                   IF (#tempRetValue <> 0) THEN
                     #LKinCtrl_OffsetContour.returnValue := #tempRetValue;
                     #LKinCtrl_OffsetContour."region" := #COFF_REGION_TYPE_RAD_COMP_LIN_CIRC;
                     #LKinCtrl_OffsetContour.subBlockNumber := 35052;
                     #LKinCtrl_OffsetContour.internalNumber := 333;
                     RETURN;
                   END_IF;



                 END_IF;

                 // Calculate end coordinate of "next" linear command
                 // Calculate orthogonal and tangential vector for next but one circular commamnd
                 #tempRetValue := "LKinCtrl_CalcCircTangOrthPathPlane"(circlePoint := #tempNextCmdIn.endPoint,
                                                                       circleCenterPoint := #tempNextButOneCmdIn.circleCenterPoint,
                                                                       pathPlane := #pathPlane,
                                                                       compDirection := #compensationDirection,
                                                                       pathChoice := #tempNextButOneCmdIn.pathChoice,
                                                                       vUnitTangentialPathPlane => #tempNextButOneCmdOut.tangentialUnitVecStart,
                                                                       vUnitOrthogonalPathPlane => #tempNextButOneCmdOut.orthogonalUnitVecStart);

                 IF (#tempRetValue <> 0) THEN
                   #LKinCtrl_OffsetContour.returnValue := #tempRetValue;
                   #LKinCtrl_OffsetContour."region" := #COFF_REGION_TYPE_RAD_COMP_LIN_CIRC;
                   #LKinCtrl_OffsetContour.subBlockNumber := 35056;
                   #LKinCtrl_OffsetContour.internalNumber := 334;
                   RETURN;
                 END_IF;


                 // Scale othogonal vector with tool radius to get orthogonal shift
                 #tempNextButOneCmdOut.orthogonalShiftStart := "LKinCtrl_VecScale"(vIn := #tempNextButOneCmdOut.orthogonalUnitVecStart,
                                                                                   factor := #toolRadius);

                 #tempNextButOneCmdOut.startPointOrthShifted := "LKinCtrl_VecAdd"(vIn1 := #tempNextCmdIn.endPoint,
                                                                                  vIn2 := #tempNextButOneCmdOut.orthogonalShiftStart);

                 // Calculate radius of circle
                 #tempNextCmdOut.circleRadius := "LKinCtrl_VecAbs"("LKinCtrl_VecSub"(vIn1 := #tempNextButOneCmdOut.startPointOrthShifted,
                                                                                                                                       vIn2 := #tempNextButOneCmdIn.circleCenterPoint));


                 // ########## Intersection point of 1st linear and 2nd circular command  ##########
                 #tempRetValue := "LKinCtrl_CalcLineCircleIntersectionPoint"(startPointLine := #tempNextCmdOut.endPointOrthShifted,
                                                                             endPointLine := #tempNextCmdOut.endPointOrthTangShifted,
                                                                             circleCenter := #tempNextButOneCmdIn.circleCenterPoint,
                                                                             circleRadius := #tempNextCmdOut.circleRadius,
                                                                             intersectionPointA => #tempPa,
                                                                             intersectionPointB => #tempPb);

                 IF (#tempRetValue <> 0) THEN
                   #LKinCtrl_OffsetContour.returnValue := #tempRetValue;
                   #LKinCtrl_OffsetContour."region" := #COFF_REGION_TYPE_RAD_COMP_LIN_CIRC;
                   #LKinCtrl_OffsetContour.subBlockNumber := 35061;
                   #LKinCtrl_OffsetContour.internalNumber := 335;
                   RETURN;
                 END_IF;

                 // Two intersection points, use the one which is closer to the circle start point
                 #tempDistance1 := "LKinCtrl_VecAbs"("LKinCtrl_VecSub"(vIn1 := #tempNextCmdOut.endPointOrthShifted, vIn2 := #tempPa));
                 #tempDistance2 := "LKinCtrl_VecAbs"("LKinCtrl_VecSub"(vIn1 := #tempNextCmdOut.endPointOrthShifted, vIn2 := #tempPb));

                 IF (#tempDistance1 < #tempDistance2) THEN
                   #tempNextCmdOut.endPoint := #tempPa;
                 ELSE
                   #tempNextCmdOut.endPoint := #tempPb;
                 END_IF;

               END_REGION
               // ############# N E X T   B U T   O N E   C M D  -  N O N E #############
             ELSE
               REGION Next but one command NONE
                 // V01.01.02 AW 2020-10-13
                 // Check if current end point is in opposite direction, e.g. small command length with big tool radius etc.
                 // Avoid reversal movement

                 // Calculate difference vector of uncompensated current and next end point
                 #tempDirectionUncompensatedVec := "LKinCtrl_VecSub"(vIn1 := #tempCurrentPoint, vIn2 := #tempNextCmdIn.endPoint);
                 #tempDirectionUncompensatedUnitVec := "LKinCtrl_VecUnit"(#tempDirectionUncompensatedVec);

                 // Calculate difference vector of compensated current and next end point
                 #tempDirectionCompensatedVec := "LKinCtrl_VecSub"(vIn1 := #tempCurrentPointRadComp, vIn2 := #tempNextCmdOut.endPoint);
                 #tempDirectionCompensatedUnitVec := "LKinCtrl_VecUnit"(#tempDirectionCompensatedVec);

                 // Calculate length between current compensated and next compensated end point
                 #tempLengthCompensatedPointDifferenceVec := "LKinCtrl_VecAbs"(#tempDirectionCompensatedVec);

                 // Check if vectors are parallel 
                 IF (((ABS(#tempDirectionUncompensatedUnitVec.x) - ABS(#tempDirectionCompensatedUnitVec.x)) < #COFF_TOLERANCE) AND
                   ((ABS(#tempDirectionUncompensatedUnitVec.y) - ABS(#tempDirectionCompensatedUnitVec.y)) < #COFF_TOLERANCE) AND
                   ((ABS(#tempDirectionUncompensatedUnitVec.z) - ABS(#tempDirectionCompensatedUnitVec.z)) < #COFF_TOLERANCE))
                 THEN
                   // Opposite direction?
                   IF ((ABS(#tempDirectionUncompensatedUnitVec.x + #tempDirectionCompensatedUnitVec.x) < #COFF_TOLERANCE) AND
                     (ABS(#tempDirectionUncompensatedUnitVec.y + #tempDirectionCompensatedUnitVec.y) < #COFF_TOLERANCE) AND
                     (ABS(#tempDirectionUncompensatedUnitVec.z + #tempDirectionCompensatedUnitVec.z) < #COFF_TOLERANCE))
                   THEN
                     // Throw error
                     #LKinCtrl_OffsetContour.returnValue := #ERR_COFF_LINEAR_CMD_AND_TOOL_RADIUS_LEAD_TO_REVERSAL;
                     #LKinCtrl_OffsetContour."region" := #COFF_REGION_TYPE_RAD_COMP_LIN_NONE;
                     #LKinCtrl_OffsetContour.subBlockNumber := 0;
                     #LKinCtrl_OffsetContour.internalNumber := 336;
                     RETURN;

                     // // Possible solution - NOT used!
                     // // Use tangential and orthogonal shift
                     // // Scale tangential vector with point difference (compensated points) to get tangential shift
                     // #tempNextCmdOut.tangentiaShiftEnd := "LKinCtrl_VecScale"(vIn := #tempNextCmdOut.tangentialUnitVecEnd,
                     //                                                          factor := #tempLengthCompensatedPointDifferenceVec);

                     // // Re-calculate orthogonal and (new) tangential shifted next target coordinate
                     // // next command end point will be equal to last command end point --> no reversal
                     // #tempNextCmdOut.endPointOrthTangShifted := "LKinCtrl_VecAdd"(vIn1 := #tempNextCmdOut.endPointOrthShifted,
                     //                                                              vIn2 := #tempNextCmdOut.tangentiaShiftEnd);

                     // // Use tangential and orthogonal shift - assign new value
                     // #tempNextCmdOut.endPoint := #tempNextCmdOut.endPointOrthTangShifted;

                   ELSE
                     // Same direction
                     ;// Nothing to do
                   END_IF;
                 ELSE
                   // V01.01.03
                   ;// Nothing to do
                 END_IF;

               END_REGION
             END_IF;

             REGION Additional plausibility check
               #tempRetValue := "LKinCtrl_CalcAngleBetweenVectors"(point1 := #tempNextCmdOut.endPoint,
                                                                   point2 := #tempNextCmdIn.endPoint,
                                                                   intersectionPoint := #tempCurrentPoint,
                                                                   angle => #tempAngle);

               IF (#tempRetValue <> 0) THEN
                 #LKinCtrl_OffsetContour.returnValue := #tempRetValue;
                 #LKinCtrl_OffsetContour."region" := #COFF_REGION_TYPE_RAD_COMP_LIN_GEN;
                 #LKinCtrl_OffsetContour.subBlockNumber := 35059;
                 #LKinCtrl_OffsetContour.internalNumber := 340;
                 RETURN;
               END_IF;

               IF (#tempAngle > #COFF_CIRC_REVERSAL_TOLERANCE_ANGLE)
               THEN
                 #LKinCtrl_OffsetContour.returnValue := #ERR_COFF_NO_SOLUTION_FOR_GIVEN_LINEAR_CMD;
                 #LKinCtrl_OffsetContour."region" := #COFF_REGION_TYPE_RAD_COMP_LIN_GEN;
                 #LKinCtrl_OffsetContour.subBlockNumber := 0;
                 #LKinCtrl_OffsetContour.internalNumber := 341;
                 RETURN;
               END_IF;

             END_REGION
           ELSE
             // Use radius compensated coordinates
             CASE #pathPlane OF
               "CP_XY":
                 #tempNextCmdOut.endPoint.x := #tempCurrentPointRadComp.x;
                 #tempNextCmdOut.endPoint.y := #tempCurrentPointRadComp.y;
                 #tempNextCmdOut.endPoint.z := #tempNextCmdOut.endPoint.z;

               "CP_XZ":
                 #tempNextCmdOut.endPoint.x := #tempCurrentPointRadComp.x;
                 #tempNextCmdOut.endPoint.y := #tempNextCmdOut.endPoint.y;
                 #tempNextCmdOut.endPoint.z := #tempCurrentPointRadComp.z;

               "CP_YZ":
                 #tempNextCmdOut.endPoint.x := #tempNextCmdOut.endPoint.x;
                 #tempNextCmdOut.endPoint.y := #tempCurrentPointRadComp.y;
                 #tempNextCmdOut.endPoint.z := #tempCurrentPointRadComp.z;
             END_CASE;
           END_IF;
         END_IF;
       END_REGION

       REGION Next command CIRCULAR
         // ############# N E X T   C M D  -  C I R C U L A R #############
         // ##############################################
         IF (#tempNextCmdOut.cmdType = "LKINCTRL_MC_MOVECIRCULARABS") THEN

           // Distinguish between different circular modes
           IF (#tempNextCmdIn.circleMode = "CM_BORDER") THEN

             // ------------ Via an intermediate point and the end point ("CircMode" = 0) ------------
             // Caluclate center point of circle with given start point, end point and intermediate point
             #tempRetValue := "LKinCtrl_CalcCircCenterByIntermediatePointAndEndPoint"(circleStartPoint := #tempCurrentPoint,
                                                                                      circleEndPoint := #tempNextCmdIn.endPoint,
                                                                                      circleIntermediatePoint := #tempNextCmdIn.circleIntermediatePoint,
                                                                                      pathPlane := #pathPlane,
                                                                                      circleCenterPoint => #tempNextCmdIn.circleCenterPoint);

             IF (#tempRetValue <> 0) THEN
               #LKinCtrl_OffsetContour.returnValue := #tempRetValue;
               #LKinCtrl_OffsetContour."region" := #COFF_REGION_TYPE_RAD_COMP_NEXT_CMD_CIRC;
               #LKinCtrl_OffsetContour.subBlockNumber := 35057;

               #LKinCtrl_OffsetContour.internalNumber := 401;
               RETURN;
             END_IF;

             // Calculate path choice
             #tempRetValue := "LKinCtrl_CalcCircPathChoiceByIntermediatePointAndEndPoint"(circleStartPoint := #tempCurrentPoint,
                                                                                          circleEndPoint := #tempNextCmdIn.endPoint,
                                                                                          circleintermediatePoint := #tempNextCmdIn.circleIntermediatePoint,
                                                                                          pathPlane := #pathPlane,
                                                                                          pathChoice => #tempNextCmdIn.pathChoice);

             IF (#tempRetValue <> 0) THEN
               #LKinCtrl_OffsetContour.returnValue := #tempRetValue;
               #LKinCtrl_OffsetContour."region" := #COFF_REGION_TYPE_RAD_COMP_NEXT_CMD_CIRC;
               #LKinCtrl_OffsetContour.subBlockNumber := 35058;
               #LKinCtrl_OffsetContour.internalNumber := 402;
               RETURN;
             END_IF;

           ELSIF (#tempNextCmdIn.circleMode = "CM_CENTER") THEN
             // ------------ Via the circle center and the angle in a main plane ("CircMode" = 1) ------------
             (* im oberen Teil!
             // "Third" coordinate is ignored by system - also ignore here!
             // Use start coordinate of circle instead
             IF (#pathPlane = "CP_XZ") THEN
               #tempNextCmdIn.circleCenterPoint.y := #tempCurrentPoint.y;
             ELSIF (#pathPlane = "CP_YZ") THEN
               #tempNextCmdIn.circleCenterPoint.x := #tempCurrentPoint.x;
             ELSIF (#pathPlane = "CP_XY") THEN
               #tempNextCmdIn.circleCenterPoint.z := #tempCurrentPoint.z;
             END_IF;*)
             ;

           ELSIF (#tempNextCmdIn.circleMode = "CM_RADIUS") THEN
             // ------------ Via the circle radius and the end point in a main plane ("CircMode" = 2) ------------
             // Calculate circle center point by given start / end point and radius and path choice
             #tempRetValue := "LKinCtrl_CalcCircCenterByRadiusAndEndPoint"(circleStartPoint := #tempCurrentPoint,
                                                                           circleEndPoint := #tempNextCmdIn.endPoint,
                                                                           pathPlane := #pathPlane,
                                                                           circleRadius := #tempNextCmdIn.circleRadius,
                                                                           pathChoice := #tempNextCmdIn.pathChoice,
                                                                           circCenterPoint => #tempNextCmdIn.circleCenterPoint);

             IF (#tempRetValue <> 0) THEN
               #LKinCtrl_OffsetContour.returnValue := #tempRetValue;
               #LKinCtrl_OffsetContour."region" := #COFF_REGION_TYPE_RAD_COMP_NEXT_CMD_CIRC;
               #LKinCtrl_OffsetContour.subBlockNumber := 35052;
               #LKinCtrl_OffsetContour.internalNumber := 403;
               RETURN;
             END_IF;

           END_IF;

           //REGION todo
           // 2019-03-07 - not necessary
           (*
           // ####
           // Calculate circle paramters
           #tempRetValue := "LKinCtrl_CalcCircTangOrthPathPlane"(circlePoint := #tempCurrentPoint,
                                                                 circleCenterPoint := #tempNextCmdIn.circleCenterPoint,
                                                                 pathPlane := #pathPlane,
                                                                 compDirection := #compensationDirection,
                                                                 pathChoice := #tempNextCmdIn.pathChoice,
                                                                 vUnitTangentialPathPlane => #tempNextCmdOut.tangentialUnitVecStart,
                                                                 vUnitOrthogonalPathPlane => #tempNextCmdOut.orthogonalUnitVecStart);

           IF (#tempRetValue <> 0) THEN
             #LKinCtrl_OffsetContour.returnValue := #tempRetValue;
             #LKinCtrl_OffsetContour."region" := #COFF_REGION_TYPE_RAD_COMP_LIN_CIRC;
             #LKinCtrl_OffsetContour.subBlockNumber := 35056;
             #LKinCtrl_OffsetContour.internalNumber := 404;
             RETURN;
           END_IF;

           // Scale othogonal vector with tool radius to get orthogonal shift
           #tempNextCmdOut.orthogonalShiftStart := "LKinCtrl_VecScale"(vIn := #tempNextCmdOut.orthogonalUnitVecStart,
                                                                       factor := #toolRadius);

           #tempNextCmdOut.startPointOrthShifted := "LKinCtrl_VecAdd"(vIn1 := #tempCurrentPoint,
                                                                      vIn2 := #tempNextCmdOut.orthogonalShiftStart);

           *)
           //END_REGION


           // #############  N E X T   B U T   O N E   C M D   #############
           // Check if next but one linear command has at least one component in path plane direction
           #tempRetValue := "LKinCtrl_CalcVecDistancePathPlane"(vectorInA := #tempNextCmdIn.endPoint,
                                                                vectorInB := #tempNextButOneCmdIn.endPoint,
                                                                pathPlane := #pathPlane,
                                                                distancePathPlane => #tempDistance1);

           IF (#tempRetValue <> 0) THEN
             #LKinCtrl_OffsetContour.returnValue := #tempRetValue;
             #LKinCtrl_OffsetContour."region" := #COFF_REGION_TYPE_RAD_COMP_CIRC_LIN;
             #LKinCtrl_OffsetContour.subBlockNumber := 35055;
             #LKinCtrl_OffsetContour.internalNumber := 405;
             RETURN;
           END_IF;

           // #############  N E X T   B U T   O N E   C M D   -  L I N E A R  #############
           // Linear command must have at least a motion in direction of path plane, otherwise treat as command none!
           IF (#tempNextButOneCmdOut.cmdType = "LKINCTRL_MC_MOVELINEARABS") AND (#tempDistance1 > 0.0) THEN

             REGION Next but one command LINEAR
               // 2nd linear command point 2 to point 3
               // Calculate tangential and orthogonal unit vector of direction (with respect to end point of circle)
               #tempRetValue := "LKinCtrl_CalcLineTangOrthPathPlane"(pathPlane := #pathPlane,
                                                                     compDirection := #compensationDirection,
                                                                     vInFirst := #tempNextButOneCmdIn.endPoint,
                                                                     vInSecond := #tempNextCmdIn.endPoint, // End point of circle
                                                                     vUnitTangentialPathPlane => #tempNextButOneCmdOut.tangentialUnitVecStart,
                                                                     vUnitOrthogonalPathPlane => #tempNextButOneCmdOut.orthogonalUnitVecStart);

               IF (#tempRetValue <> 0) THEN
                 #LKinCtrl_OffsetContour.returnValue := #tempRetValue;
                 #LKinCtrl_OffsetContour."region" := #COFF_REGION_TYPE_RAD_COMP_CIRC_LIN;
                 #LKinCtrl_OffsetContour.subBlockNumber := 35055;
                 #LKinCtrl_OffsetContour.internalNumber := 406;
                 RETURN;
               END_IF;

               // Scale othogonal vector with tool radius to get orthogonal shift
               #tempNextButOneCmdOut.orthogonalShiftStart := "LKinCtrl_VecScale"(vIn := #tempNextButOneCmdOut.orthogonalUnitVecStart,
                                                                                 factor := #toolRadius);

               // Scale tangential vector with tool radius to get tangential shift
               #tempNextButOneCmdOut.tangentiaShiftStart := "LKinCtrl_VecScale"(vIn := #tempNextButOneCmdOut.tangentialUnitVecStart,
                                                                                factor := #toolRadius);

               // Calculate orthogonal shifted next target coordinate
               #tempNextButOneCmdOut.startPointOrthShifted := "LKinCtrl_VecAdd"(vIn1 := #tempNextCmdIn.endPoint, // Start coordinate next but one command
                                                                                vIn2 := #tempNextButOneCmdOut.orthogonalShiftStart);

               // Calculate orthogonal and tangential shifted next target coordinate
               #tempNextButOneCmdOut.startPointOrthTangShifted := "LKinCtrl_VecAdd"(vIn1 := #tempNextButOneCmdOut.startPointOrthShifted,
                                                                                    vIn2 := #tempNextButOneCmdOut.tangentiaShiftStart);

               // ########## Intersection point of 1st circular and 2nd linear command  ##########
               // Change center point to same level with start point
               IF (#tempNextCmdIn.circleMode = "CM_BORDER") THEN
                 // ------------ Via an intermediate point and the end point ("CircMode" = 0) ------------
                 // 3D circle possible

                 // Bring circle parameter to the same level as current point
                 #tempNextCmdEndPointLevelled := #tempNextCmdIn.endPoint;
                 #tempNextCmdIntermediatePointLevelled := #tempNextCmdIn.circleIntermediatePoint;


                 // Bring coordinates to same level as current point
                 #tempNextCmdStartPointOrhtShiftLevelled := #tempCurrentPointRadComp;// #tempNextCmdOut.startPointOrthShifted;
                 #tempNextButOneStartPointOrthShiftedLevelled := #tempNextButOneCmdOut.startPointOrthShifted;
                 #tempNextButOneCmdStartPointOrthTangShiftedLevelled := #tempNextButOneCmdOut.startPointOrthTangShifted;

                 // Level parameters (third coordinate) with current point
                 CASE #pathPlane OF
                   "CP_XZ":
                     #tempNextCmdEndPointLevelled.y := #tempCurrentPoint.y;
                     #tempNextCmdIntermediatePointLevelled.y := #tempCurrentPoint.y;
                     #tempNextCmdStartPointOrhtShiftLevelled.y := #tempCurrentPoint.y;
                     #tempNextButOneStartPointOrthShiftedLevelled.y := #tempCurrentPoint.y;
                     #tempNextButOneCmdStartPointOrthTangShiftedLevelled.y := #tempCurrentPoint.y;

                   "CP_YZ":
                     #tempNextCmdEndPointLevelled.x := #tempCurrentPoint.x;
                     #tempNextCmdIntermediatePointLevelled.x := #tempCurrentPoint.x;
                     #tempNextCmdStartPointOrhtShiftLevelled.x := #tempCurrentPoint.x;
                     #tempNextButOneStartPointOrthShiftedLevelled.x := #tempCurrentPoint.x;
                     #tempNextButOneCmdStartPointOrthTangShiftedLevelled.x := #tempCurrentPoint.x;

                   "CP_XY":
                     #tempNextCmdEndPointLevelled.z := #tempCurrentPoint.z;
                     #tempNextCmdIntermediatePointLevelled.z := #tempCurrentPoint.z;
                     #tempNextCmdStartPointOrhtShiftLevelled.z := #tempCurrentPoint.z;
                     #tempNextButOneStartPointOrthShiftedLevelled.z := #tempCurrentPoint.z;
                     #tempNextButOneCmdStartPointOrthTangShiftedLevelled.z := #tempCurrentPoint.z;
                   ELSE
                     #LKinCtrl_OffsetContour.returnValue := #ERR_COFF_INTERNAL;
                     #LKinCtrl_OffsetContour."region" := #COFF_REGION_TYPE_RAD_COMP_CIRC_LIN;
                     #LKinCtrl_OffsetContour.internalNumber := 407;
                     RETURN;
                 END_CASE;

                 // Calculate new levelled circle center point
                 #tempRetValue := "LKinCtrl_CalcCircCenterByIntermediatePointAndEndPoint"(circleStartPoint := #tempCurrentPoint,
                                                                                          circleEndPoint := #tempNextCmdEndPointLevelled,
                                                                                          circleIntermediatePoint := #tempNextCmdIntermediatePointLevelled,
                                                                                          pathPlane := #pathPlane,
                                                                                          circleCenterPoint => #tempNextCmdOut.circleCenterPoint); // levelled

                 IF (#tempRetValue <> 0) THEN
                   #LKinCtrl_OffsetContour.returnValue := #tempRetValue;
                   #LKinCtrl_OffsetContour."region" := #COFF_REGION_TYPE_RAD_COMP_NEXT_CMD_CIRC;
                   #LKinCtrl_OffsetContour.subBlockNumber := 35057;
                   #LKinCtrl_OffsetContour.internalNumber := 408;
                   RETURN;
                 END_IF;

                 // Calculate modified radius - levelled
                 #tempNextCmdOut.circleRadius := "LKinCtrl_VecAbs"("LKinCtrl_VecSub"(vIn1 := #tempNextCmdStartPointOrhtShiftLevelled,
                                                                                     vIn2 := #tempNextCmdOut.circleCenterPoint));




                 #tempRetValue := "LKinCtrl_CalcLineCircleIntersectionPoint"(startPointLine := #tempNextButOneStartPointOrthShiftedLevelled,
                                                                             endPointLine := #tempNextButOneCmdStartPointOrthTangShiftedLevelled,
                                                                             circleCenter := #tempNextCmdOut.circleCenterPoint,
                                                                             circleRadius := #tempNextCmdOut.circleRadius,
                                                                             intersectionPointA => #tempPa,
                                                                             intersectionPointB => #tempPb);

                 // Relevel intersection point
                 CASE #pathPlane OF
                   "CP_XZ":
                     #tempPa.y := #tempNextCmdIn.endPoint.y;
                     #tempPb.y := #tempNextCmdIn.endPoint.y;

                   "CP_YZ":
                     #tempPa.x := #tempNextCmdIn.endPoint.x;
                     #tempPb.x := #tempNextCmdIn.endPoint.x;

                   "CP_XY":
                     #tempPa.z := #tempNextCmdIn.endPoint.z;
                     #tempPb.z := #tempNextCmdIn.endPoint.z;
                   ELSE
                     #LKinCtrl_OffsetContour.returnValue := #ERR_COFF_INTERNAL;
                     #LKinCtrl_OffsetContour."region" := #COFF_REGION_TYPE_RAD_COMP_CIRC_LIN;
                     #LKinCtrl_OffsetContour.internalNumber := 409;
                     RETURN;
                 END_CASE;

               ELSE
                 // 2D circle
                 // Calculate modified radius
                 #tempNextCmdOut.circleRadius := "LKinCtrl_VecAbs"("LKinCtrl_VecSub"(vIn1 := #tempCurrentPointRadComp,//#tempNextCmdOut.startPointOrthShifted,
                                                                                     vIn2 := #tempNextCmdIn.circleCenterPoint));

                 #tempRetValue := "LKinCtrl_CalcLineCircleIntersectionPoint"(startPointLine := #tempNextButOneCmdOut.startPointOrthShifted,
                                                                             endPointLine := #tempNextButOneCmdOut.startPointOrthTangShifted,
                                                                             circleCenter := #tempNextCmdIn.circleCenterPoint,
                                                                             circleRadius := #tempNextCmdOut.circleRadius,
                                                                             intersectionPointA => #tempPa,
                                                                             intersectionPointB => #tempPb);


               END_IF;


               IF (#tempRetValue <> 0) THEN
                 #LKinCtrl_OffsetContour.returnValue := #tempRetValue;
                 #LKinCtrl_OffsetContour."region" := #COFF_REGION_TYPE_RAD_COMP_CIRC_LIN;
                 #LKinCtrl_OffsetContour.subBlockNumber := 35061;
                 #LKinCtrl_OffsetContour.internalNumber := 410;
                 RETURN;
               END_IF;

               // Two intersection points, use the one which is closer to the circle end point
               #tempDistance1 := "LKinCtrl_VecAbs"("LKinCtrl_VecSub"(vIn1 := #tempNextCmdIn.endPoint, vIn2 := #tempPa));
               #tempDistance2 := "LKinCtrl_VecAbs"("LKinCtrl_VecSub"(vIn1 := #tempNextCmdIn.endPoint, vIn2 := #tempPb));

               IF (#tempDistance1 < #tempDistance2) THEN
                 #tempNextCmdOut.endPoint := #tempPa;
               ELSE
                 #tempNextCmdOut.endPoint := #tempPb;
               END_IF;

             END_REGION
             // #############  N E X T   B U T   O N E   C M D   -  C I R C U L A R #############
           ELSIF (#tempNextButOneCmdOut.cmdType = "LKINCTRL_MC_MOVECIRCULARABS") THEN
             REGION Next but one command CIRCULAR
               // Distinguish between different circular modes
               IF (#tempNextButOneCmdIn.circleMode = "CM_BORDER") THEN
                 // ------------ Via an intermediate point and the end point ("CircMode" = 0) ------------

                 // Caluclate center point of circle with given start point, end point and intermediate point
                 #tempRetValue := "LKinCtrl_CalcCircCenterByIntermediatePointAndEndPoint"(circleStartPoint := #tempNextCmdIn.endPoint,
                                                                                          circleEndPoint := #tempNextButOneCmdIn.endPoint,
                                                                                          circleIntermediatePoint := #tempNextButOneCmdIn.circleIntermediatePoint,
                                                                                          pathPlane := #pathPlane,
                                                                                          circleCenterPoint => #tempNextButOneCmdIn.circleCenterPoint);

                 IF (#tempRetValue <> 0) THEN
                   #LKinCtrl_OffsetContour.returnValue := #tempRetValue;
                   #LKinCtrl_OffsetContour."region" := #COFF_REGION_TYPE_RAD_COMP_CIRC_CIRC;
                   #LKinCtrl_OffsetContour.subBlockNumber := 35057;
                   #LKinCtrl_OffsetContour.internalNumber := 430;
                   RETURN;
                 END_IF;

                 // Calculate path choice
                 #tempRetValue := "LKinCtrl_CalcCircPathChoiceByIntermediatePointAndEndPoint"(circleStartPoint := #tempNextCmdIn.endPoint,
                                                                                              circleEndPoint := #tempNextButOneCmdIn.endPoint,
                                                                                              circleintermediatePoint := #tempNextButOneCmdIn.circleIntermediatePoint,
                                                                                              pathPlane := #pathPlane,
                                                                                              pathChoice => #tempNextButOneCmdIn.pathChoice);

                 IF (#tempRetValue <> 0) THEN
                   #LKinCtrl_OffsetContour.returnValue := #tempRetValue;
                   #LKinCtrl_OffsetContour."region" := #COFF_REGION_TYPE_RAD_COMP_CIRC_CIRC;
                   #LKinCtrl_OffsetContour.subBlockNumber := 35058;
                   #LKinCtrl_OffsetContour.internalNumber := 431;
                   RETURN;
                 END_IF;

               ELSIF (#tempNextButOneCmdIn.circleMode = "CM_CENTER") THEN
                 // ------------ Via the circle center and the angle in a main plane ("CircMode" = 1) ------------

                 // "Third" coordinate is ignored by system - also ignore here!
                 // Use start coordinate of circle instead
                 IF (#pathPlane = "CP_XZ") THEN
                   #tempNextButOneCmdIn.circleCenterPoint.y := #tempNextCmdIn.endPoint.y;
                 ELSIF (#pathPlane = "CP_YZ") THEN
                   #tempNextButOneCmdIn.circleCenterPoint.x := #tempNextCmdIn.endPoint.x;
                 ELSIF (#pathPlane = "CP_XY") THEN
                   #tempNextButOneCmdIn.circleCenterPoint.z := #tempNextCmdIn.endPoint.z;
                 END_IF;

                 // Calculte correct circle end point - parameter not mandatory (and therefore probably not correct)
                 #tempRetValue := "LKinCtrl_CalcCircEndPointWithGivenCenterAndAngle"(circleStartPoint := #tempNextCmdIn.endPoint,
                                                                                     circleCenterPoint := #tempNextButOneCmdIn.circleCenterPoint,
                                                                                     pathPlane := #pathPlane,
                                                                                     pathChoice := #tempNextButOneCmdIn.pathChoice,
                                                                                     angle := #tempNextButOneCmdIn.circleAngle,
                                                                                     endPoint => #tempNextButOneCmdIn.endPoint);

                 IF (#tempRetValue <> 0) THEN
                   #LKinCtrl_OffsetContour.returnValue := #tempRetValue;
                   #LKinCtrl_OffsetContour."region" := #COFF_REGION_TYPE_RAD_COMP_CIRC_CIRC;
                   #LKinCtrl_OffsetContour.subBlockNumber := 35053;
                   #LKinCtrl_OffsetContour.internalNumber := 432;
                   RETURN;
                 END_IF;

               ELSIF (#tempNextButOneCmdIn.circleMode = "CM_RADIUS") THEN
                 // ------------ Via the circle radius and the end point in a main plane ("CircMode" = 2) ------------
                 #tempRetValue := "LKinCtrl_CalcCircCenterByRadiusAndEndPoint"(circleStartPoint := #tempNextCmdIn.endPoint,
                                                                               circleEndPoint := #tempNextButOneCmdIn.endPoint,
                                                                               pathPlane := #pathPlane,
                                                                               circleRadius := #tempNextButOneCmdIn.circleRadius,
                                                                               pathChoice := #tempNextButOneCmdIn.pathChoice,
                                                                               circCenterPoint => #tempNextButOneCmdIn.circleCenterPoint);

                 IF (#tempRetValue <> 0) THEN
                   #LKinCtrl_OffsetContour.returnValue := #tempRetValue;
                   #LKinCtrl_OffsetContour."region" := #COFF_REGION_TYPE_RAD_COMP_CIRC_CIRC;
                   #LKinCtrl_OffsetContour.subBlockNumber := 35052;
                   #LKinCtrl_OffsetContour.internalNumber := 433;
                   RETURN;
                 END_IF;

               END_IF;

               // Take care of next circular command
               #tempRetValue := "LKinCtrl_CalcCircTangOrthPathPlane"(circlePoint := #tempNextCmdIn.endPoint,
                                                                     circleCenterPoint := #tempNextButOneCmdIn.circleCenterPoint,
                                                                     pathPlane := #pathPlane,
                                                                     compDirection := #compensationDirection,
                                                                     pathChoice := #tempNextButOneCmdIn.pathChoice,
                                                                     vUnitTangentialPathPlane => #tempNextButOneCmdOut.tangentialUnitVecStart,
                                                                     vUnitOrthogonalPathPlane => #tempNextButOneCmdOut.orthogonalUnitVecStart);

               IF (#tempRetValue <> 0) THEN
                 #LKinCtrl_OffsetContour.returnValue := #tempRetValue;
                 #LKinCtrl_OffsetContour."region" := #COFF_REGION_TYPE_RAD_COMP_CIRC_CIRC;
                 #LKinCtrl_OffsetContour.subBlockNumber := 35056;
                 #LKinCtrl_OffsetContour.internalNumber := 434;
                 RETURN;
               END_IF;

               // Scale othogonal vector with tool radius to get orthogonal shift
               #tempNextButOneCmdOut.orthogonalShiftStart := "LKinCtrl_VecScale"(vIn := #tempNextButOneCmdOut.orthogonalUnitVecStart,
                                                                                 factor := #toolRadius);


               #tempNextButOneCmdOut.startPointOrthShifted := "LKinCtrl_VecAdd"(vIn1 := #tempNextCmdIn.endPoint,
                                                                                vIn2 := #tempNextButOneCmdOut.orthogonalShiftStart);

               // ########## Intersection point of 1st circular and 2nd circular command  ##########

               IF (#tempNextCmdIn.circleMode = "CM_BORDER") THEN
                 // ------------ Via an intermediate point and the end point ("CircMode" = 0) ------------
                 // 3D circle possible
                 // 
                 // Bring coordinates and parameters to same level as current point
                 #tempNextCmdStartPointOrhtShiftLevelled := #tempCurrentPointRadComp; //#tempNextCmdOut.startPointOrthShifted;
                 #tempNextCmdOut.circleCenterPoint := #tempNextCmdIn.circleCenterPoint;

                 // Level parameters (third coordinate) with current point
                 CASE #pathPlane OF
                   "CP_XZ":
                     #tempNextCmdStartPointOrhtShiftLevelled.y := #tempCurrentPoint.y;
                     #tempNextCmdOut.circleCenterPoint.y := #tempCurrentPoint.y;

                   "CP_YZ":
                     #tempNextCmdStartPointOrhtShiftLevelled.x := #tempCurrentPoint.x;
                     #tempNextCmdOut.circleCenterPoint.x := #tempCurrentPoint.x;

                   "CP_XY":
                     #tempNextCmdStartPointOrhtShiftLevelled.z := #tempCurrentPoint.z;
                     #tempNextCmdOut.circleCenterPoint.z := #tempCurrentPoint.z;
                   ELSE
                     #LKinCtrl_OffsetContour.returnValue := #ERR_COFF_INTERNAL;
                     #LKinCtrl_OffsetContour."region" := #COFF_REGION_TYPE_RAD_COMP_CIRC_CIRC;
                     #LKinCtrl_OffsetContour.internalNumber := 435;
                     RETURN;
                 END_CASE;

                 // Calculate radius of shifted 1st circle - levelled
                 #tempNextCmdOut.circleRadius := "LKinCtrl_VecAbs"("LKinCtrl_VecSub"(vIn1 := #tempNextCmdStartPointOrhtShiftLevelled,
                                                                                     vIn2 := #tempNextCmdOut.circleCenterPoint));
               ELSE
                 #tempNextCmdOut.circleCenterPoint := #tempNextCmdIn.circleCenterPoint;
                 // Calculate radius of shifted 1st circle
                 #tempNextCmdOut.circleRadius := "LKinCtrl_VecAbs"("LKinCtrl_VecSub"(vIn1 := #tempCurrentPointRadComp,
                                                                                     vIn2 := #tempNextCmdOut.circleCenterPoint));
               END_IF;

               IF (#tempNextButOneCmdIn.circleMode = "CM_BORDER") THEN
                 // ------------ Via an intermediate point and the end point ("CircMode" = 0) ------------
                 // 3D circle possible
                 // 
                 // Bring coordinates and parameters to same level as current point
                 #tempNextButOneStartPointOrthShiftedLevelled := #tempNextButOneCmdOut.startPointOrthShifted;
                 #tempNextButOneCmdOut.circleCenterPoint := #tempNextButOneCmdIn.circleCenterPoint;

                 // Level parameters (third coordinate) with current point
                 CASE #pathPlane OF
                   "CP_XZ":
                     #tempNextButOneStartPointOrthShiftedLevelled.y := #tempCurrentPoint.y;
                     #tempNextButOneCmdOut.circleCenterPoint.y := #tempCurrentPoint.y;

                   "CP_YZ":
                     #tempNextButOneStartPointOrthShiftedLevelled.x := #tempCurrentPoint.x;
                     #tempNextButOneCmdOut.circleCenterPoint.x := #tempCurrentPoint.x;

                   "CP_XY":
                     #tempNextButOneStartPointOrthShiftedLevelled.z := #tempCurrentPoint.z;
                     #tempNextButOneCmdOut.circleCenterPoint.z := #tempCurrentPoint.z;
                   ELSE
                     #LKinCtrl_OffsetContour.returnValue := #ERR_COFF_INTERNAL;
                     #LKinCtrl_OffsetContour."region" := #COFF_REGION_TYPE_RAD_COMP_CIRC_CIRC;
                     #LKinCtrl_OffsetContour.internalNumber := 435;
                     RETURN;
                 END_CASE;
                 // Calculate radius of shifted 2nd circle - levelled
                 #tempNextButOneCmdOut.circleRadius := "LKinCtrl_VecAbs"("LKinCtrl_VecSub"(vIn1 := #tempNextButOneStartPointOrthShiftedLevelled,
                                                                                           vIn2 := #tempNextButOneCmdOut.circleCenterPoint));
               ELSE
                 #tempNextButOneCmdOut.circleCenterPoint := #tempNextButOneCmdIn.circleCenterPoint;

                 // Calculate radius of shifted 2nd circle
                 // preliminary
                 #tempNextButOneCmdOut.circleRadius := "LKinCtrl_VecAbs"("LKinCtrl_VecSub"(vIn1 := #tempNextButOneCmdOut.startPointOrthShifted,
                                                                                           vIn2 := #tempNextButOneCmdOut.circleCenterPoint));
               END_IF;

               // Intersection point of 1st and 2nd circle
               #tempRetValue := "LKinCtrl_CalcCircleCircleIntersectionPoint"(circleCenterPoint1 := #tempNextCmdOut.circleCenterPoint,
                                                                             circleCenterPoint2 := #tempNextButOneCmdOut.circleCenterPoint,
                                                                             circleRadius1 := #tempNextCmdOut.circleRadius,
                                                                             circleRadius2 := #tempNextButOneCmdOut.circleRadius,
                                                                             pathPlane := #pathPlane,
                                                                             intersectionPointA => #tempPa,
                                                                             intersectionPointB => #tempPb);
               IF (#tempRetValue <> 0) THEN
                 // V01.00.01
                 IF (#tempRetValue = #ERR_COFF_CIRCLE_CENTERS_EQUAL) THEN
                   // Circles are equal - use modified start point of following circle instead
                   #tempPa := #tempNextButOneCmdOut.startPointOrthShifted;
                   #tempPb := #tempNextButOneCmdOut.startPointOrthShifted;
                 ELSE
                   #LKinCtrl_OffsetContour.returnValue := #tempRetValue;
                   #LKinCtrl_OffsetContour."region" := #COFF_REGION_TYPE_RAD_COMP_CIRC_CIRC;
                   #LKinCtrl_OffsetContour.subBlockNumber := 35062;
                   #LKinCtrl_OffsetContour.internalNumber := 437;
                   RETURN;
                 END_IF;
               END_IF;

               IF (#tempNextCmdIn.circleMode = "CM_BORDER") THEN
                 // ------------ Via an intermediate point and the end point ("CircMode" = 0) ------------
                 // 3D circle possible
                 // Relevel intersection point
                 CASE #pathPlane OF
                   "CP_XZ":
                     #tempPa.y := #tempNextCmdIn.endPoint.y;
                     #tempPb.y := #tempNextCmdIn.endPoint.y;

                   "CP_YZ":
                     #tempPa.x := #tempNextCmdIn.endPoint.x;
                     #tempPb.x := #tempNextCmdIn.endPoint.x;

                   "CP_XY":
                     #tempPa.z := #tempNextCmdIn.endPoint.z;
                     #tempPb.z := #tempNextCmdIn.endPoint.z;
                   ELSE
                     #LKinCtrl_OffsetContour.returnValue := #ERR_COFF_INTERNAL;
                     #LKinCtrl_OffsetContour."region" := #COFF_REGION_TYPE_RAD_COMP_CIRC_LIN;
                     #LKinCtrl_OffsetContour.internalNumber := 436;
                     RETURN;
                 END_CASE;
               END_IF;

               // Two intersection points, use the one which is closer to the circle end point
               #tempDistance1 := "LKinCtrl_VecAbs"("LKinCtrl_VecSub"(vIn1 := #tempNextCmdIn.endPoint, vIn2 := #tempPa));
               #tempDistance2 := "LKinCtrl_VecAbs"("LKinCtrl_VecSub"(vIn1 := #tempNextCmdIn.endPoint, vIn2 := #tempPb));

               IF (#tempDistance1 < #tempDistance2) THEN
                 #tempNextCmdOut.endPoint := #tempPa;
               ELSE
                 #tempNextCmdOut.endPoint := #tempPb;
               END_IF;

             END_REGION
             // ############# N E X T   B U T   O N E   C M D  -  N O N E #############
           ELSE
             REGION Next but one command NONE
               // Output next but one coordinates - in case it's the last one
               #tempNextButOneCmdOut.endPoint := #tempNextButOneCmdOut.endPointOrthShifted;

               // Calculate end point for circle (orthogonal shifted)
               #tempRetValue := "LKinCtrl_CalcCircTangOrthPathPlane"(circlePoint := #tempNextCmdIn.endPoint,
                                                                     circleCenterPoint := #tempNextCmdIn.circleCenterPoint,
                                                                     pathPlane := #pathPlane,
                                                                     compDirection := #compensationDirection,
                                                                     pathChoice := #tempNextCmdIn.pathChoice,
                                                                     vUnitTangentialPathPlane => #tempNextCmdOut.tangentialUnitVecEnd,
                                                                     vUnitOrthogonalPathPlane => #tempNextCmdOut.orthogonalUnitVecEnd);

               IF (#tempRetValue <> 0) THEN
                 #LKinCtrl_OffsetContour.returnValue := #tempRetValue;
                 #LKinCtrl_OffsetContour."region" := #COFF_REGION_TYPE_RAD_COMP_CIRC_NONE;
                 #LKinCtrl_OffsetContour.subBlockNumber := 35056;
                 #LKinCtrl_OffsetContour.internalNumber := 450;
                 RETURN;
               END_IF;

               // Scale othogonal vector with tool radius to get orthogonal shift
               #tempNextCmdOut.orthogonalShiftEnd := "LKinCtrl_VecScale"(vIn := #tempNextCmdOut.orthogonalUnitVecEnd,
                                                                         factor := #toolRadius);


               #tempNextCmdOut.endPoint := "LKinCtrl_VecAdd"(vIn1 := #tempNextCmdIn.endPoint,
                                                             vIn2 := #tempNextCmdOut.orthogonalShiftEnd);
               (*
               // Distinguish between different circular modes
               IF (#tempNextCmdIn.circleMode = "CM_BORDER") THEN
                 // ------------ Via an intermediate point and the end point ("CircMode" = 0) ------------

                 // Calculate end point for circle mode 0 by given mode 0
                 #tempRetValue := "LKinCtrl_CalcCircTangOrthPathPlane"(circlePoint := #tempNextCmdIn.endPoint,
                                                                       circleCenterPoint := #tempNextCmdIn.circleCenterPoint,
                                                                       pathPlane := #pathPlane,
                                                                       compDirection := #compensationDirection,
                                                                       pathChoice := #tempNextCmdIn.pathChoice,
                                                                       vUnitTangentialPathPlane => #tempNextCmdOut.tangentialUnitVecEnd,
                                                                       vUnitOrthogonalPathPlane => #tempNextCmdOut.orthogonalUnitVecEnd);

                 IF (#tempRetValue <> 0) THEN
                   #LKinCtrl_OffsetContour.returnValue := #tempRetValue;
                   #LKinCtrl_OffsetContour."region" := #COFF_REGION_TYPE_RAD_COMP_CIRC_NONE;
                   #LKinCtrl_OffsetContour.subBlockNumber := 35056;
                   #LKinCtrl_OffsetContour.internalNumber := 450;
                   RETURN;
                 END_IF;

                 // Scale othogonal vector with tool radius to get orthogonal shift
                 #tempNextCmdOut.orthogonalShiftEnd := "LKinCtrl_VecScale"(vIn := #tempNextCmdOut.orthogonalUnitVecEnd,
                                                                           factor := #toolRadius);
